VERSION : 0.1
   VAR_INPUT
      "BUFFER STATE" : Int;
      "ITEMS COUNT" : Int;
      "DOWN ELEVATOR LEFT SENSOR" : Bool;
      "BRIDGE SENSOR 1" : Bool;
      "BRIDGE SENSOR 2" : Bool;
   END_VAR
   VAR_OUTPUT
      "Z3-1 BRIDGE" : Bool;
      "Z3-2 BRIDGE" : Bool;
      "Z3-3 BRIDGE" : Bool;
   END_VAR
   VAR
      F_TRIG_Instance : F_TRIG;
      "DOWN SENSOR TRIG" : Bool;
      "BRIDGE SENSOR 1 TRIG" : Bool;
      "BRIDGE SENSOR 2 TRIG" : Bool;
      F_TRIG_BS1 : F_TRIG;
      F_TRIG_BS2 : F_TRIG;
   END_VAR
BEGIN
   #F_TRIG_Instance(CLK := #"DOWN ELEVATOR LEFT SENSOR",
                    Q => #"DOWN SENSOR TRIG");
   #F_TRIG_BS1(CLK := #"BRIDGE SENSOR 1",
               Q => #"BRIDGE SENSOR 1 TRIG");
   #F_TRIG_BS2(CLK := #"BRIDGE SENSOR 2",
               Q => #"BRIDGE SENSOR 2 TRIG");
   CASE #"ITEMS COUNT" OF
       1..2:
           #"Z3-3 BRIDGE" := 1;
           #"Z3-2 BRIDGE" := 0;
           #"Z3-3 BRIDGE" := 0;

           IF #"DOWN SENSOR TRIG" THEN
               #"Z3-3 BRIDGE" := 0;
               #"Z3-2 BRIDGE" := 0;
               #"Z3-3 BRIDGE" := 0;


           END_IF;
       3..4:
           #"Z3-3 BRIDGE" := 1;
           #"Z3-2 BRIDGE" := 1;
           #"Z3-3 BRIDGE" := 0;

           IF #"BRIDGE SENSOR 2 TRIG" AND #"DOWN SENSOR TRIG" THEN
               #"Z3-3 BRIDGE" := 0;
               #"Z3-2 BRIDGE" := 0;
               #"Z3-3 BRIDGE" := 0;

           END_IF;
       5..6:
           #"Z3-3 BRIDGE" := 1;
           #"Z3-2 BRIDGE" := 1;
           #"Z3-3 BRIDGE":=1;

           IF #"BRIDGE SENSOR 2 TRIG" AND #"DOWN SENSOR TRIG" AND #"BRIDGE SENSOR 1 TRIG" THEN
               #"Z3-3 BRIDGE" := 0;
               #"Z3-2 BRIDGE" := 0;
               #"Z3-3 BRIDGE" := 0;

           END_IF;
       ELSE 
           #"Z3-3 BRIDGE" := 0;
           #"Z3-2 BRIDGE" := 0;
           #"Z3-3 BRIDGE" := 0;

   END_CASE;
END_FUNCTION_BLOCK

FUNCTION_BLOCK "ZONE 3 ELEVATORS LOGIC"   // FB11, SCL
{ S7_Optimized_Access := 'TRUE' }
VERSION : 0.1
   VAR_INPUT
      "BUFFER STATE" : Int;
   END_VAR
   VAR_OUTPUT
      "UP ELEVATOR" : Bool;
      "DOWN ELEVATOR" : Bool;
   END_VAR
BEGIN
   IF #"BUFFER STATE" = 10 OR #"BUFFER STATE" = 33 OR #"BUFFER STATE" = 36 OR #"BUFFER STATE" = 39 THEN
       #"UP ELEVATOR" := 1;
       #"DOWN ELEVATOR" := 0;
   ELSIF #"BUFFER STATE" = 70 OR #"BUFFER STATE"=50 THEN
       #"UP ELEVATOR" := 0;
       #"DOWN ELEVATOR" := 1;
   ELSE
       #"UP ELEVATOR" := 0;
       #"DOWN ELEVATOR" := 0;
   END_IF;
END_FUNCTION_BLOCK

FUNCTION_BLOCK "ZONE 3 BRIDGE CONVS LOGIC"   // FB12, SCL
{ S7_Optimized_Access := 'TRUE' }
VERSION : 0.1
   VAR_INPUT
      "BUFFER STATE" : Int;
      "BRIDGE SENSOR 1" : Bool;
      "BRIDGE SENSOR 2" : Bool;
      "UP ELEVATOR SENSOR RIGHT" : Bool;
      "DOWN ELEVATOR LEFT SENSOR" : Bool;
      "ITEMS COUNT" : Int;
   END_VAR
   VAR_OUTPUT
      "Z3-1 BRIDGE" : Bool;
      "Z3-2 BRIDGE" : Bool;
      "Z3-3 BRIDGE" : Bool;
      "STATE 50 DONE" : Bool;
      "STATE 30 DONE" : Bool;
   END_VAR
   VAR
      "bridge sensor 1 set" : Bool;
      "bridge sensor 2 set" : Bool;
      "elevator sensor set" : Bool;
   END_VAR
BEGIN
   IF #"BUFFER STATE" = 33 THEN
       #"Z3-1 BRIDGE" := 1;
       #"Z3-2 BRIDGE" := 1;
       #"Z3-3 BRIDGE" := 1;
       IF #"BRIDGE SENSOR 2" THEN
           #"Z3-1 BRIDGE" := 0;
           #"Z3-2 BRIDGE" := 0;
           #"Z3-3 BRIDGE" := 0;
           #"STATE 30 DONE" := 1;
       END_IF;
   ELSIF #"BUFFER STATE" = 36 THEN
       #"Z3-1 BRIDGE" := 1;
       #"Z3-2 BRIDGE" := 1;
       #"Z3-3 BRIDGE" := 0;
       IF #"BRIDGE SENSOR 1" THEN
           #"Z3-1 BRIDGE" := 0;
           #"Z3-2 BRIDGE" := 0;
           #"Z3-3 BRIDGE" := 0;
           #"STATE 30 DONE" := 1;
       END_IF;
   ELSIF #"BUFFER STATE" = 39 THEN
       #"Z3-1 BRIDGE" := 1;
       #"Z3-2 BRIDGE" := 0;
       #"Z3-3 BRIDGE" := 0;
       IF #"UP ELEVATOR SENSOR RIGHT" THEN
           #"Z3-1 BRIDGE" := 0;
           #"Z3-2 BRIDGE" := 0;
           #"Z3-3 BRIDGE" := 0;
           #"STATE 30 DONE" := 1;
       END_IF;
   ELSIF #"BUFFER STATE" = 50 THEN
       CASE #"ITEMS COUNT" OF
           0..1:(*

        modified the item count to be less by one because at the cycle scan it is degreesed before it reads the current value
   *)
               #"Z3-3 BRIDGE" := 1;
               #"Z3-2 BRIDGE" := 0;
               #"Z3-1 BRIDGE" := 0;

               IF #"DOWN ELEVATOR LEFT SENSOR" THEN
                   #"Z3-3 BRIDGE" := 0;
                   #"Z3-2 BRIDGE" := 0;
                   #"Z3-1 BRIDGE" := 0;
                   #"STATE 50 DONE" := 1;

               END_IF;
           2..3:
               #"Z3-3 BRIDGE" := 1;
               #"Z3-2 BRIDGE" := 1;
               #"Z3-1 BRIDGE" := 0;

               IF #"BRIDGE SENSOR 2" THEN
                   #"bridge sensor 2 set" := 1;
               END_IF;
               IF #"DOWN ELEVATOR LEFT SENSOR" THEN
                   #"elevator sensor set" := 1;
               END_IF;
               IF #"bridge sensor 2 set" AND #"elevator sensor set" THEN
                   #"Z3-3 BRIDGE" := 0;
                   #"Z3-2 BRIDGE" := 0;
                   #"Z3-1 BRIDGE" := 0;
                   #"STATE 50 DONE" := 1;
                   #"bridge sensor 2 set" :=0;
                   #"elevator sensor set" :=0;
               END_IF;
           4..6:
               #"Z3-3 BRIDGE" := 1;
               #"Z3-2 BRIDGE" := 1;
               #"Z3-1 BRIDGE" := 1;

               IF #"BRIDGE SENSOR 2" THEN
                   #"bridge sensor 2 set" := 1;
               END_IF;
               IF #"DOWN ELEVATOR LEFT SENSOR" THEN
                   #"elevator sensor set" := 1;
               END_IF;
               IF #"BRIDGE SENSOR 1" THEN
                   #"bridge sensor 1 set" := 1;
               END_IF;
               IF #"bridge sensor 1 set" AND #"bridge sensor 2 set" AND #"elevator sensor set" THEN
                   #"Z3-3 BRIDGE" := 0;
                   #"Z3-2 BRIDGE" := 0;
                   #"Z3-1 BRIDGE" := 0;
                   #"STATE 50 DONE" := 1;
                   #"bridge sensor 2 set" := 0;
                   #"elevator sensor set" := 0;
                   #"bridge sensor 1 set" := 0;
               END_IF;
           ELSE
               #"Z3-3 BRIDGE" := 0;
               #"Z3-2 BRIDGE" := 0;
               #"Z3-1 BRIDGE" := 0;

       END_CASE;
   ELSE
       #"Z3-1 BRIDGE" := 0;
       #"Z3-2 BRIDGE" := 0;
       #"Z3-3 BRIDGE" := 0;
       #"STATE 30 DONE" := 0;
       #"STATE 50 DONE" := 0;
   END_IF;
END_FUNCTION_BLOCK

(* ===== HMI "HMI_RT_1" =====
system functions are stored by id; their names below are inferred from use
connection "HMI_Connection_1": ETHERNET, SMART_S7_1200_OMS

HMI tags "Default tag table"
   "Tag_ScreenNumber" : UInt, internal
   "DB_RackMemory_In_Production" : Int = PLC DB_RackMemory.In_Production, 1 s
   "ZONE-3 BUFFER_A_DB_BUFFER_ITEMS_COUNT_CV" : Int = PLC "ZONE-3 BUFFER_A_DB".BUFFER_ITEMS_COUNT.CV, 1 s
   "Zone_3_FB_DB_ZONE-3 BUFFER B_BUFFER_ITEMS_COUNT_CV" : Int = PLC Zone_3_FB_DB."ZONE-3 BUFFER B".BUFFER_ITEMS_COUNT.CV, 1 s
   "DB_RackMemory_SpacesOccupied" : Int = PLC DB_RackMemory.SpacesOccupied, 1 s
   "DB_HMI_Z3 BUFFER A STATUS" : Int = PLC DB_HMI."Z3 BUFFER A STATUS", 1 s
   "DB_HMI_Z1 STATUS" : Int = PLC DB_HMI."Z1 STATUS", 1 s
   "DB_HMI_Z2 STATUS" : Int = PLC DB_HMI."Z2 STATUS", 1 s
   "DB_HMI_Z3 BUFFER B STATUS" : Int = PLC DB_HMI."Z3 BUFFER B STATUS", 1 s
   "DB_HMI_Z3 ASSEMPLER STATUS" : Int = PLC DB_HMI."Z3 ASSEMPLER STATUS", 1 s
   "DB_HMI_Z5 STATUS" : Int = PLC DB_HMI."Z5 STATUS", 1 s
   "DB_HMI_Z4 UPPER STATUS" : Int = PLC DB_HMI."Z4 UPPER STATUS", 1 s
   "DB_HMI_Z4 LOWER STATUS" : Int = PLC DB_HMI."Z4 LOWER STATUS", 1 s
   "DB_HMI_FACTORY STATUS" : Int = PLC DB_HMI."FACTORY STATUS", 1 s
   "DB_RackMemory_QUANTITY TO RETRIEVE" : Int = PLC DB_RackMemory."QUANTITY TO RETRIEVE", 1 s
   "DB_RackMemory_TOTAL ORDERS" : Int = PLC DB_RackMemory."TOTAL ORDERS", 1 s
   "DB_RackMemory_TOTAL DLIEVERED" : Int = PLC DB_RackMemory."TOTAL DLIEVERED", 1 s
   "DB_RackMemory_REQUIRED QUANTITY" : Int = PLC DB_RackMemory."REQUIRED QUANTITY", 1 s
   "DB_HMI_CREATE ORDER" : Bool = PLC DB_HMI."CREATE ORDER", 1 s
   "DB_HMI_CANCEL ORDER" : Bool = PLC DB_HMI."CANCEL ORDER", 1 s
   "DB_RackMemory_FREE SPACES" : Int = PLC DB_RackMemory."FREE SPACES", 1 s
   "DB_RackMemory_Rack{1}_occupied" : Bool = PLC DB_RackMemory.Rack[1].occupied, 1 s
   "DB_RackMemory_Rack{2}_occupied" : Bool = PLC DB_RackMemory.Rack[2].occupied, 1 s
   "DB_RackMemory_Rack{3}_occupied" : Bool = PLC DB_RackMemory.Rack[3].occupied, 1 s
   "DB_RackMemory_Rack{4}_occupied" : Bool = PLC DB_RackMemory.Rack[4].occupied, 1 s
   "DB_RackMemory_Rack{5}_occupied" : Bool = PLC DB_RackMemory.Rack[5].occupied, 1 s
   "DB_RackMemory_Rack{6}_occupied" : Bool = PLC DB_RackMemory.Rack[6].occupied, 1 s
   "DB_RackMemory_Rack{7}_occupied" : Bool = PLC DB_RackMemory.Rack[7].occupied, 1 s
   "DB_RackMemory_Rack{8}_occupied" : Bool = PLC DB_RackMemory.Rack[8].occupied, 1 s
   "DB_RackMemory_Rack{9}_occupied" : Bool = PLC DB_RackMemory.Rack[9].occupied, 1 s
   "DB_RackMemory_Rack{10}_occupied" : Bool = PLC DB_RackMemory.Rack[10].occupied, 1 s
   "DB_RackMemory_Rack{11}_occupied" : Bool = PLC DB_RackMemory.Rack[11].occupied, 1 s
   "DB_RackMemory_Rack{12}_occupied" : Bool = PLC DB_RackMemory.Rack[12].occupied, 1 s
   "DB_RackMemory_Rack{13}_occupied" : Bool = PLC DB_RackMemory.Rack[13].occupied, 1 s
   "DB_RackMemory_Rack{14}_occupied" : Bool = PLC DB_RackMemory.Rack[14].occupied, 1 s
   "DB_RackMemory_Rack{15}_occupied" : Bool = PLC DB_RackMemory.Rack[15].occupied, 1 s
   "DB_RackMemory_Rack{16}_occupied" : Bool = PLC DB_RackMemory.Rack[16].occupied, 1 s
   "DB_RackMemory_Rack{17}_occupied" : Bool = PLC DB_RackMemory.Rack[17].occupied, 1 s
   "DB_RackMemory_Rack{18}_occupied" : Bool = PLC DB_RackMemory.Rack[18].occupied, 1 s
   "DB_RackMemory_Rack{19}_occupied" : Bool = PLC DB_RackMemory.Rack[19].occupied, 1 s
   "DB_RackMemory_Rack{20}_occupied" : Bool = PLC DB_RackMemory.Rack[20].occupied, 1 s
   "DB_RackMemory_Rack{21}_occupied" : Bool = PLC DB_RackMemory.Rack[21].occupied, 1 s
   "DB_RackMemory_Rack{22}_occupied" : Bool = PLC DB_RackMemory.Rack[22].occupied, 1 s
   "DB_RackMemory_Rack{23}_occupied" : Bool = PLC DB_RackMemory.Rack[23].occupied, 1 s
   "DB_RackMemory_Rack{24}_occupied" : Bool = PLC DB_RackMemory.Rack[24].occupied, 1 s
   "DB_RackMemory_Rack{25}_occupied" : Bool = PLC DB_RackMemory.Rack[25].occupied, 1 s
   "DB_RackMemory_Rack{26}_occupied" : Bool = PLC DB_RackMemory.Rack[26].occupied, 1 s
   "DB_RackMemory_Rack{27}_occupied" : Bool = PLC DB_RackMemory.Rack[27].occupied, 1 s
   "DB_RackMemory_Rack{28}_occupied" : Bool = PLC DB_RackMemory.Rack[28].occupied, 1 s
   "DB_RackMemory_Rack{29}_occupied" : Bool = PLC DB_RackMemory.Rack[29].occupied, 1 s
   "DB_RackMemory_Rack{30}_occupied" : Bool = PLC DB_RackMemory.Rack[30].occupied, 1 s
   "DB_RackMemory_Rack{31}_occupied" : Bool = PLC DB_RackMemory.Rack[31].occupied, 1 s
   "DB_RackMemory_Rack{32}_occupied" : Bool = PLC DB_RackMemory.Rack[32].occupied, 1 s
   "DB_RackMemory_Rack{33}_occupied" : Bool = PLC DB_RackMemory.Rack[33].occupied, 1 s
   "DB_RackMemory_Rack{34}_occupied" : Bool = PLC DB_RackMemory.Rack[34].occupied, 1 s
   "DB_RackMemory_Rack{35}_occupied" : Bool = PLC DB_RackMemory.Rack[35].occupied, 1 s
   "DB_RackMemory_Rack{36}_occupied" : Bool = PLC DB_RackMemory.Rack[36].occupied, 1 s
   "DB_RackMemory_Rack{37}_occupied" : Bool = PLC DB_RackMemory.Rack[37].occupied, 1 s
   "DB_RackMemory_Rack{38}_occupied" : Bool = PLC DB_RackMemory.Rack[38].occupied, 1 s
   "DB_RackMemory_Rack{39}_occupied" : Bool = PLC DB_RackMemory.Rack[39].occupied, 1 s
   "DB_RackMemory_Rack{40}_occupied" : Bool = PLC DB_RackMemory.Rack[40].occupied, 1 s
   "DB_RackMemory_Rack{41}_occupied" : Bool = PLC DB_RackMemory.Rack[41].occupied, 1 s
   "DB_RackMemory_Rack{42}_occupied" : Bool = PLC DB_RackMemory.Rack[42].occupied, 1 s
   "DB_RackMemory_Rack{43}_occupied" : Bool = PLC DB_RackMemory.Rack[43].occupied, 1 s
   "DB_RackMemory_Rack{44}_occupied" : Bool = PLC DB_RackMemory.Rack[44].occupied, 1 s
   "DB_RackMemory_Rack{45}_occupied" : Bool = PLC DB_RackMemory.Rack[45].occupied, 1 s
   "DB_RackMemory_Rack{46}_occupied" : Bool = PLC DB_RackMemory.Rack[46].occupied, 1 s
   "DB_RackMemory_Rack{47}_occupied" : Bool = PLC DB_RackMemory.Rack[47].occupied, 1 s
   "DB_RackMemory_Rack{48}_occupied" : Bool = PLC DB_RackMemory.Rack[48].occupied, 1 s
   "DB_RackMemory_Rack{49}_occupied" : Bool = PLC DB_RackMemory.Rack[49].occupied, 1 s
   "DB_RackMemory_Rack{50}_occupied" : Bool = PLC DB_RackMemory.Rack[50].occupied, 1 s
   "DB_RackMemory_Rack{51}_occupied" : Bool = PLC DB_RackMemory.Rack[51].occupied, 1 s
   "DB_RackMemory_Rack{52}_occupied" : Bool = PLC DB_RackMemory.Rack[52].occupied, 1 s
   "DB_RackMemory_Rack{53}_occupied" : Bool = PLC DB_RackMemory.Rack[53].occupied, 1 s
   "DB_RackMemory_Rack{54}_occupied" : Bool = PLC DB_RackMemory.Rack[54].occupied, 1 s
   "DB_RackMemory_Rack{55}_occupied" : Bool = PLC DB_RackMemory.Rack[55].occupied, 1 s
   "DB_RackMemory_Rack{56}_occupied" : Bool = PLC DB_RackMemory.Rack[56].occupied, 1 s
   "DB_RackMemory_Rack{57}_occupied" : Bool = PLC DB_RackMemory.Rack[57].occupied, 1 s
   "DB_RackMemory_Rack{58}_occupied" : Bool = PLC DB_RackMemory.Rack[58].occupied, 1 s
   "DB_RackMemory_Rack{59}_occupied" : Bool = PLC DB_RackMemory.Rack[59].occupied, 1 s
   "DB_RackMemory_Rack{60}_occupied" : Bool = PLC DB_RackMemory.Rack[60].occupied, 1 s
   "DB_RackMemory_Rack{61}_occupied" : Bool = PLC DB_RackMemory.Rack[61].occupied, 1 s
   "DB_RackMemory_Rack{62}_occupied" : Bool = PLC DB_RackMemory.Rack[62].occupied, 1 s
   "DB_RackMemory_Rack{63}_occupied" : Bool = PLC DB_RackMemory.Rack[63].occupied, 1 s
   "DB_RackMemory_Rack{64}_occupied" : Bool = PLC DB_RackMemory.Rack[64].occupied, 1 s
   "DB_RackMemory_Rack{65}_occupied" : Bool = PLC DB_RackMemory.Rack[65].occupied, 1 s
   "DB_RackMemory_Rack{66}_occupied" : Bool = PLC DB_RackMemory.Rack[66].occupied, 1 s
   "DB_RackMemory_Rack{67}_occupied" : Bool = PLC DB_RackMemory.Rack[67].occupied, 1 s
   "DB_RackMemory_Rack{68}_occupied" : Bool = PLC DB_RackMemory.Rack[68].occupied, 1 s
   "DB_RackMemory_Rack{69}_occupied" : Bool = PLC DB_RackMemory.Rack[69].occupied, 1 s
   "DB_RackMemory_Rack{70}_occupied" : Bool = PLC DB_RackMemory.Rack[70].occupied, 1 s
   "DB_RackMemory_Rack{71}_occupied" : Bool = PLC DB_RackMemory.Rack[71].occupied, 1 s
   "DB_RackMemory_Rack{72}_occupied" : Bool = PLC DB_RackMemory.Rack[72].occupied, 1 s
   "DB_RackMemory_Rack{73}_occupied" : Bool = PLC DB_RackMemory.Rack[73].occupied, 1 s
   "DB_RackMemory_Rack{74}_occupied" : Bool = PLC DB_RackMemory.Rack[74].occupied, 1 s
   "DB_RackMemory_Rack{75}_occupied" : Bool = PLC DB_RackMemory.Rack[75].occupied, 1 s
   "DB_RackMemory_Rack{76}_occupied" : Bool = PLC DB_RackMemory.Rack[76].occupied, 1 s
   "DB_RackMemory_Rack{77}_occupied" : Bool = PLC DB_RackMemory.Rack[77].occupied, 1 s
   "DB_RackMemory_Rack{78}_occupied" : Bool = PLC DB_RackMemory.Rack[78].occupied, 1 s
   "DB_RackMemory_Rack{79}_occupied" : Bool = PLC DB_RackMemory.Rack[79].occupied, 1 s
   "DB_RackMemory_Rack{80}_occupied" : Bool = PLC DB_RackMemory.Rack[80].occupied, 1 s
   "DB_RackMemory_Rack{81}_occupied" : Bool = PLC DB_RackMemory.Rack[81].occupied, 1 s
   "DB_RackMemory_Rack{82}_occupied" : Bool = PLC DB_RackMemory.Rack[82].occupied, 1 s
   "DB_RackMemory_Rack{83}_occupied" : Bool = PLC DB_RackMemory.Rack[83].occupied, 1 s
   "DB_RackMemory_Rack{84}_occupied" : Bool = PLC DB_RackMemory.Rack[84].occupied, 1 s
   "DB_RackMemory_Rack{85}_occupied" : Bool = PLC DB_RackMemory.Rack[85].occupied, 1 s
   "DB_RackMemory_Rack{86}_occupied" : Bool = PLC DB_RackMemory.Rack[86].occupied, 1 s
   "DB_RackMemory_Rack{87}_occupied" : Bool = PLC DB_RackMemory.Rack[87].occupied, 1 s
   "DB_RackMemory_Rack{88}_occupied" : Bool = PLC DB_RackMemory.Rack[88].occupied, 1 s
   "DB_RackMemory_Rack{89}_occupied" : Bool = PLC DB_RackMemory.Rack[89].occupied, 1 s
   "DB_RackMemory_Rack{90}_occupied" : Bool = PLC DB_RackMemory.Rack[90].occupied, 1 s
   "DB_RackMemory_Rack{91}_occupied" : Bool = PLC DB_RackMemory.Rack[91].occupied, 1 s
   "DB_RackMemory_Rack{92}_occupied" : Bool = PLC DB_RackMemory.Rack[92].occupied, 1 s
   "DB_RackMemory_Rack{93}_occupied" : Bool = PLC DB_RackMemory.Rack[93].occupied, 1 s
   "DB_RackMemory_Rack{94}_occupied" : Bool = PLC DB_RackMemory.Rack[94].occupied, 1 s
   "DB_RackMemory_Rack{95}_occupied" : Bool = PLC DB_RackMemory.Rack[95].occupied, 1 s
   "DB_RackMemory_Rack{96}_occupied" : Bool = PLC DB_RackMemory.Rack[96].occupied, 1 s
   "DB_RackMemory_Rack{97}_occupied" : Bool = PLC DB_RackMemory.Rack[97].occupied, 1 s
   "DB_RackMemory_Rack{98}_occupied" : Bool = PLC DB_RackMemory.Rack[98].occupied, 1 s
   "DB_RackMemory_Rack{99}_occupied" : Bool = PLC DB_RackMemory.Rack[99].occupied, 1 s
   "DB_RackMemory_Rack{100}_occupied" : Bool = PLC DB_RackMemory.Rack[100].occupied, 1 s
   "DB_RackMemory_Rack{101}_occupied" : Bool = PLC DB_RackMemory.Rack[101].occupied, 1 s
   "DB_RackMemory_Rack{102}_occupied" : Bool = PLC DB_RackMemory.Rack[102].occupied, 1 s
   "DB_RackMemory_Rack{103}_occupied" : Bool = PLC DB_RackMemory.Rack[103].occupied, 1 s
   "DB_RackMemory_Rack{104}_occupied" : Bool = PLC DB_RackMemory.Rack[104].occupied, 1 s
   "DB_RackMemory_Rack{105}_occupied" : Bool = PLC DB_RackMemory.Rack[105].occupied, 1 s
   "DB_RackMemory_Rack{106}_occupied" : Bool = PLC DB_RackMemory.Rack[106].occupied, 1 s
   "DB_RackMemory_Rack{107}_occupied" : Bool = PLC DB_RackMemory.Rack[107].occupied, 1 s
   "DB_RackMemory_Rack{108}_occupied" : Bool = PLC DB_RackMemory.Rack[108].occupied, 1 s
   "DB_HMI_CRANE TARGET" : Int = PLC DB_HMI."CRANE TARGET", 1 s
   "DB_HMI_CRANE SIDE" : Int = PLC DB_HMI."CRANE SIDE", 1 s
   "DB_HMI_ASSEMPLER X" : Real = PLC DB_HMI."ASSEMPLER X", 1 s
   "DB_HMI_ASSEMPLER Z" : Real = PLC DB_HMI."ASSEMPLER Z", 1 s
   "DB_RackMemory_ReckMemoryReset" : Bool = PLC DB_RackMemory.ReckMemoryReset, 1 s
   "DB_RackMemory_InProductionReset" : Bool = PLC DB_RackMemory.InProductionReset, 1 s
   "DB_HMI_CRANE LIFT" : Bool = PLC DB_HMI."CRANE LIFT", 1 s
   "DB_HMI_CRANE LEFT" : Bool = PLC DB_HMI."CRANE LEFT", 1 s
   "DB_HMI_CRANE RIGHT" : Bool = PLC DB_HMI."CRANE RIGHT", 1 s
   "DB_HMI_ASSEMPLER ROT CW" : Bool = PLC DB_HMI."ASSEMPLER ROT CW", 1 s
   "DB_HMI_ASSEMPLER ROT CCW" : Bool = PLC DB_HMI."ASSEMPLER ROT CCW", 1 s
   "DB_HMI_ASSEMPLER GRAB" : Bool = PLC DB_HMI."ASSEMPLER GRAB", 1 s
   "DB_RackMemory_RETRIEVE" : Bool = PLC DB_RackMemory.RETRIEVE, 1 s
   "CURRENT USER" : WString[254] AT %DB1.DBX0.0
   "DB_HMI_MAINTENANCE MODE" : Bool = PLC DB_HMI."MAINTENANCE MODE", 1 s

HMI tags "Alarm tag table"
   "Alarm_Trigger" : Word = PLC Alarm_trigger AT %MW100, 1 s

discrete alarms
   1: 'Emergency button is pressed', class Errors, trigger "Alarm_Trigger" bit 0
   2: 'MACHINE A HAS AN ERROR AND STOPPED WORKING', class Errors, trigger "Alarm_Trigger" bit 1
   3: 'MACHINE B HAS AN ERROR AND STOPPED WORKING', class Errors, trigger "Alarm_Trigger" bit 2
   4: 'BUFFER A HAS A PROBLEM AND STOPPED RESPONDING', class Errors, trigger "Alarm_Trigger" bit 3
   5: 'BUFFER B HAS A PROBLEM AND STOPPED WORKING', class Errors, trigger "Alarm_Trigger" bit 4
   6: 'ASSEMPLER HAS A PROBLEM AND STOPPED RESPONDING', class Errors, trigger "Alarm_Trigger" bit 5
   7: 'PALLETIZER HAS A PROBLEM AND STOPPED RESPONDING', class Errors, trigger "Alarm_Trigger" bit 6
   8: 'CRANE HAS A PROBLEM AND STOPPED RESPONDING', class Errors, trigger "Alarm_Trigger" bit 7

Template "Template_1" 800x480
   Button "Template_Button" at 714,429 size 71x50; TextOff 'Text'
   Button "Template_Button_1" at 614,429 size 71x50; TextOff 'Text'
   Button "Template_Button_2" at 514,429 size 71x50; TextOff 'Text'
   Button "Template_Button_3" at 414,429 size 71x50; TextOff 'Text'
   Button "Template_Button_4" at 314,429 size 71x50; TextOff 'Text'
   Button "Template_Button_5" at 214,429 size 71x50; TextOff 'Text'
   Button "Template_Button_6" at 114,429 size 71x50; TextOff 'Text'
   Button "Template_Button_7" at 14,429 size 71x50; TextOff 'Text'
   SymbolicIOField "Symbolic_IO_Field_Screen" at 93,9 size 600x33; TextOff '0'; TextOn '1'; TextList "TextList_ScreenNames"
      ProcessValue <- "Tag_ScreenNumber"
      on Change: ActivateScreenByNumber("Tag_ScreenNumber", 0)
   DateTimeField "HmiScreenItemData" at 695,25 size 105x25
   DateTimeField "HmiScreenItemData_1" at 695,0 size 105x25
   GraphicView "Logo" at 0,0 size 91x51; Picture "Logo of HMI_1"

screen "Production" 800x480
   Button "Button_12" at 69,415 size 163x52; TextOff 'Overview'
      on Release: ActivateScreen("Overview", 0)
   Button "Button_13" at 238,415 size 163x52; TextOff 'Warehouse'
      on Release: ActivateScreen("Warehouse", 0)
   Button "Button_14" at 408,415 size 163x52; TextOff 'Alarms'
      on Release: ActivateScreen("Alarms", 0)
   Button "Button_15" at 578,415 size 163x52; TextOff 'Maintenance'; Authorization "Maintenance"
      on Release: ActivateScreen("Maintenance", 0)
   TextField "Text field_1" at 310,0 size 180x44; Text 'Production'
   TextField "Text field_2" at 12,130 size 86x23; Text 'Quantity :'
   IOField "I/O field_1" at 124,121 size 96x32; Authorization "Operate"; FormatPattern 99
      ProcessValue <- "DB_RackMemory_QUANTITY TO RETRIEVE"
   Button "Button_1" at 65,221 size 96x32; TextOff 'Order'; Authorization "Operate"
      on Press: SetBit("DB_RackMemory_RETRIEVE")
   TextField "Text field_3" at 128,307 size 97x23; Text 'In Storage:'
   TextField "Text field_4" at 381,307 size 164x23; Text 'In Production lines:'
   IOField "I/O field_2" at 255,298 size 96x32; FormatPattern 999
      ProcessValue <- "DB_RackMemory_SpacesOccupied"
   IOField "I/O field_3" at 575,298 size 96x32; FormatPattern 99
      ProcessValue <- "DB_RackMemory_In_Production"
   TextField "Text field_5" at 27,70 size 163x33; Text 'Create Order:'
   TextField "Text field_6" at 312,70 size 175x33; Text 'Current Order:'
   TextField "Text field_7" at 247,130 size 161x23; Text 'Required Products:'
   TextField "Text field_8" at 240,183 size 174x23; Text 'Products Remaining:'
   TextField "Text field_9" at 610,70 size 124x33; Text 'Summary:'
   TextField "Text field_10" at 558,130 size 113x23; Text 'Total Orders:'
   TextField "Text field_11" at 537,183 size 147x23; Text 'Total Delievered:'
   Button "Button_2" at 352,221 size 96x32; TextOff 'Cancel'; Authorization "Operate"
      on Press: SetBit("DB_HMI_CANCEL ORDER")
      on Release: ResetBit("DB_HMI_CANCEL ORDER")
   IOField "I/O field_4" at 425,121 size 96x32; FormatPattern 99
      ProcessValue <- "DB_RackMemory_REQUIRED QUANTITY"
   IOField "I/O field_5" at 425,174 size 96x32; FormatPattern 99
      ProcessValue <- "DB_RackMemory_QUANTITY TO RETRIEVE"
   IOField "I/O field_6" at 690,121 size 96x32; FormatPattern 999
      ProcessValue <- "DB_RackMemory_TOTAL ORDERS"
   IOField "I/O field_7" at 690,174 size 96x32; FormatPattern 999
      ProcessValue <- "DB_RackMemory_TOTAL DLIEVERED"
   Button "Button_3" at 11,10 size 96x32; TextOff 'LOG IN'
      on Release: function_f41c6f6c("CURRENT USER")
      on Press: function_a2a04561()
   Button "Button_4" at 126,8 size 96x32; TextOff 'LOG OUT'
      on Press: function_f23ef4c9(); SetTag("CURRENT USER", '""')
   IOField "I/O field_13" at 685,3 size 106x32; FormatPattern ??????????????????????????????????????????????????????????????????????
      ProcessValue <- "CURRENT USER"
   TextField "Text field_12" at 542,8 size 140x23; Text 'CURRENT USER:'

screen "Warehouse" 800x480
   Rectangle "Rectangle_1" at 698,216 size 20x20
      Appearance <- "DB_RackMemory_Rack{1}_occupied"
   Rectangle "Rectangle_2" at 678,216 size 20x20
      Appearance <- "DB_RackMemory_Rack{2}_occupied"
   Rectangle "Rectangle_3" at 658,216 size 20x20
      Appearance <- "DB_RackMemory_Rack{3}_occupied"
   Rectangle "Rectangle_4" at 638,216 size 20x20
      Appearance <- "DB_RackMemory_Rack{4}_occupied"
   Rectangle "Rectangle_5" at 618,216 size 20x20
      Appearance <- "DB_RackMemory_Rack{5}_occupied"
   Rectangle "Rectangle_6" at 598,216 size 20x20
      Appearance <- "DB_RackMemory_Rack{6}_occupied"
   Rectangle "Rectangle_7" at 578,216 size 20x20
      Appearance <- "DB_RackMemory_Rack{7}_occupied"
   Rectangle "Rectangle_8" at 558,216 size 20x20
      Appearance <- "DB_RackMemory_Rack{8}_occupied"
   Rectangle "Rectangle_9" at 538,216 size 20x20
      Appearance <- "DB_RackMemory_Rack{9}_occupied"
   Rectangle "Rectangle_10" at 698,196 size 20x20
      Appearance <- "DB_RackMemory_Rack{10}_occupied"
   Rectangle "Rectangle_11" at 678,196 size 20x20
      Appearance <- "DB_RackMemory_Rack{11}_occupied"
   Rectangle "Rectangle_12" at 658,196 size 20x20
      Appearance <- "DB_RackMemory_Rack{12}_occupied"
   Rectangle "Rectangle_13" at 638,196 size 20x20
      Appearance <- "DB_RackMemory_Rack{13}_occupied"
   Rectangle "Rectangle_14" at 618,196 size 20x20
      Appearance <- "DB_RackMemory_Rack{14}_occupied"
   Rectangle "Rectangle_15" at 598,196 size 20x20
      Appearance <- "DB_RackMemory_Rack{15}_occupied"
   Rectangle "Rectangle_16" at 578,196 size 20x20
      Appearance <- "DB_RackMemory_Rack{16}_occupied"
   Rectangle "Rectangle_17" at 558,196 size 20x20
      Appearance <- "DB_RackMemory_Rack{17}_occupied"
   Rectangle "Rectangle_18" at 538,196 size 20x20
      Appearance <- "DB_RackMemory_Rack{18}_occupied"
   Rectangle "Rectangle_19" at 698,176 size 20x20
      Appearance <- "DB_RackMemory_Rack{19}_occupied"
   Rectangle "Rectangle_20" at 678,176 size 20x20
      Appearance <- "DB_RackMemory_Rack{20}_occupied"
   Rectangle "Rectangle_21" at 658,176 size 20x20
      Appearance <- "DB_RackMemory_Rack{21}_occupied"
   Rectangle "Rectangle_22" at 638,176 size 20x20
      Appearance <- "DB_RackMemory_Rack{22}_occupied"
   Rectangle "Rectangle_23" at 618,176 size 20x20
      Appearance <- "DB_RackMemory_Rack{23}_occupied"
   Rectangle "Rectangle_24" at 598,176 size 20x20
      Appearance <- "DB_RackMemory_Rack{24}_occupied"
   Rectangle "Rectangle_25" at 578,176 size 20x20
      Appearance <- "DB_RackMemory_Rack{25}_occupied"
   Rectangle "Rectangle_26" at 558,176 size 20x20
      Appearance <- "DB_RackMemory_Rack{26}_occupied"
   Rectangle "Rectangle_27" at 538,176 size 20x20
      Appearance <- "DB_RackMemory_Rack{27}_occupied"
   Rectangle "Rectangle_28" at 698,156 size 20x20
      Appearance <- "DB_RackMemory_Rack{28}_occupied"
   Rectangle "Rectangle_29" at 678,156 size 20x20
      Appearance <- "DB_RackMemory_Rack{29}_occupied"
   Rectangle "Rectangle_30" at 658,156 size 20x20
      Appearance <- "DB_RackMemory_Rack{30}_occupied"
   Rectangle "Rectangle_31" at 638,156 size 20x20
      Appearance <- "DB_RackMemory_Rack{31}_occupied"
   Rectangle "Rectangle_32" at 618,156 size 20x20
      Appearance <- "DB_RackMemory_Rack{32}_occupied"
   Rectangle "Rectangle_33" at 598,156 size 20x20
      Appearance <- "DB_RackMemory_Rack{33}_occupied"
   Rectangle "Rectangle_34" at 578,156 size 20x20
      Appearance <- "DB_RackMemory_Rack{34}_occupied"
   Rectangle "Rectangle_35" at 558,156 size 20x20
      Appearance <- "DB_RackMemory_Rack{35}_occupied"
   Rectangle "Rectangle_36" at 538,156 size 20x20
      Appearance <- "DB_RackMemory_Rack{36}_occupied"
   Rectangle "Rectangle_37" at 698,136 size 20x20
      Appearance <- "DB_RackMemory_Rack{37}_occupied"
   Rectangle "Rectangle_38" at 678,136 size 20x20
      Appearance <- "DB_RackMemory_Rack{38}_occupied"
   Rectangle "Rectangle_39" at 658,136 size 20x20
      Appearance <- "DB_RackMemory_Rack{39}_occupied"
   Rectangle "Rectangle_40" at 638,136 size 20x20
      Appearance <- "DB_RackMemory_Rack{40}_occupied"
   Rectangle "Rectangle_41" at 618,136 size 20x20
      Appearance <- "DB_RackMemory_Rack{41}_occupied"
   Rectangle "Rectangle_42" at 598,136 size 20x20
      Appearance <- "DB_RackMemory_Rack{42}_occupied"
   Rectangle "Rectangle_43" at 578,136 size 20x20
      Appearance <- "DB_RackMemory_Rack{43}_occupied"
   Rectangle "Rectangle_44" at 558,136 size 20x20
      Appearance <- "DB_RackMemory_Rack{44}_occupied"
   Rectangle "Rectangle_45" at 538,136 size 20x20
      Appearance <- "DB_RackMemory_Rack{45}_occupied"
   Rectangle "Rectangle_46" at 698,116 size 20x20
      Appearance <- "DB_RackMemory_Rack{46}_occupied"
   Rectangle "Rectangle_47" at 678,116 size 20x20
      Appearance <- "DB_RackMemory_Rack{47}_occupied"
   Rectangle "Rectangle_48" at 658,116 size 20x20
      Appearance <- "DB_RackMemory_Rack{48}_occupied"
   Rectangle "Rectangle_49" at 638,116 size 20x20
      Appearance <- "DB_RackMemory_Rack{49}_occupied"
   Rectangle "Rectangle_50" at 618,116 size 20x20
      Appearance <- "DB_RackMemory_Rack{50}_occupied"
   Rectangle "Rectangle_51" at 598,116 size 20x20
      Appearance <- "DB_RackMemory_Rack{51}_occupied"
   Rectangle "Rectangle_52" at 578,116 size 20x20
      Appearance <- "DB_RackMemory_Rack{52}_occupied"
   Rectangle "Rectangle_53" at 558,116 size 20x20
      Appearance <- "DB_RackMemory_Rack{53}_occupied"
   Rectangle "Rectangle_54" at 538,116 size 20x20
      Appearance <- "DB_RackMemory_Rack{54}_occupied"
   Rectangle "Rectangle_69" at 142,196 size 20x20
      Appearance <- "DB_RackMemory_Rack{69}_occupied"
   Rectangle "Rectangle_55" at 242,216 size 20x20
      Appearance <- "DB_RackMemory_Rack{55}_occupied"
   Rectangle "Rectangle_56" at 222,216 size 20x20
      Appearance <- "DB_RackMemory_Rack{56}_occupied"
   Rectangle "Rectangle_57" at 202,216 size 20x20
      Appearance <- "DB_RackMemory_Rack{57}_occupied"
   Rectangle "Rectangle_58" at 182,216 size 20x20
      Appearance <- "DB_RackMemory_Rack{58}_occupied"
   Rectangle "Rectangle_59" at 162,216 size 20x20
      Appearance <- "DB_RackMemory_Rack{59}_occupied"
   Rectangle "Rectangle_60" at 142,216 size 20x20
      Appearance <- "DB_RackMemory_Rack{60}_occupied"
   Rectangle "Rectangle_61" at 122,216 size 20x20
      Appearance <- "DB_RackMemory_Rack{61}_occupied"
   Rectangle "Rectangle_62" at 102,216 size 20x20
      Appearance <- "DB_RackMemory_Rack{62}_occupied"
   Rectangle "Rectangle_63" at 82,216 size 20x20
      Appearance <- "DB_RackMemory_Rack{63}_occupied"
   Rectangle "Rectangle_64" at 242,196 size 20x20
      Appearance <- "DB_RackMemory_Rack{64}_occupied"
   Rectangle "Rectangle_65" at 222,196 size 20x20
      Appearance <- "DB_RackMemory_Rack{65}_occupied"
   Rectangle "Rectangle_66" at 202,196 size 20x20
      Appearance <- "DB_RackMemory_Rack{66}_occupied"
   Rectangle "Rectangle_67" at 182,196 size 20x20
      Appearance <- "DB_RackMemory_Rack{67}_occupied"
   Rectangle "Rectangle_68" at 162,196 size 20x20
      Appearance <- "DB_RackMemory_Rack{68}_occupied"
   Rectangle "Rectangle_70" at 122,196 size 20x20
      Appearance <- "DB_RackMemory_Rack{70}_occupied"
   Rectangle "Rectangle_71" at 102,196 size 20x20
      Appearance <- "DB_RackMemory_Rack{71}_occupied"
   Rectangle "Rectangle_72" at 82,196 size 20x20
      Appearance <- "DB_RackMemory_Rack{72}_occupied"
   Rectangle "Rectangle_73" at 242,176 size 20x20
      Appearance <- "DB_RackMemory_Rack{73}_occupied"
   Rectangle "Rectangle_74" at 222,176 size 20x20
      Appearance <- "DB_RackMemory_Rack{74}_occupied"
   Rectangle "Rectangle_75" at 202,176 size 20x20
      Appearance <- "DB_RackMemory_Rack{75}_occupied"
   Rectangle "Rectangle_76" at 182,176 size 20x20
      Appearance <- "DB_RackMemory_Rack{76}_occupied"
   Rectangle "Rectangle_77" at 162,176 size 20x20
      Appearance <- "DB_RackMemory_Rack{77}_occupied"
   Rectangle "Rectangle_78" at 142,176 size 20x20
      Appearance <- "DB_RackMemory_Rack{78}_occupied"
   Rectangle "Rectangle_79" at 122,176 size 20x20
      Appearance <- "DB_RackMemory_Rack{79}_occupied"
   Rectangle "Rectangle_80" at 102,176 size 20x20
      Appearance <- "DB_RackMemory_Rack{80}_occupied"
   Rectangle "Rectangle_81" at 82,176 size 20x20
      Appearance <- "DB_RackMemory_Rack{81}_occupied"
   Rectangle "Rectangle_82" at 242,156 size 20x20
      Appearance <- "DB_RackMemory_Rack{82}_occupied"
   Rectangle "Rectangle_83" at 222,156 size 20x20
      Appearance <- "DB_RackMemory_Rack{83}_occupied"
   Rectangle "Rectangle_84" at 202,156 size 20x20
      Appearance <- "DB_RackMemory_Rack{84}_occupied"
   Rectangle "Rectangle_85" at 182,156 size 20x20
      Appearance <- "DB_RackMemory_Rack{85}_occupied"
   Rectangle "Rectangle_86" at 162,156 size 20x20
      Appearance <- "DB_RackMemory_Rack{86}_occupied"
   Rectangle "Rectangle_87" at 142,156 size 20x20
      Appearance <- "DB_RackMemory_Rack{87}_occupied"
   Rectangle "Rectangle_88" at 122,156 size 20x20
      Appearance <- "DB_RackMemory_Rack{88}_occupied"
   Rectangle "Rectangle_89" at 102,156 size 20x20
      Appearance <- "DB_RackMemory_Rack{89}_occupied"
   Rectangle "Rectangle_90" at 82,156 size 20x20
      Appearance <- "DB_RackMemory_Rack{90}_occupied"
   Rectangle "Rectangle_91" at 242,136 size 20x20
      Appearance <- "DB_RackMemory_Rack{91}_occupied"
   Rectangle "Rectangle_92" at 222,136 size 20x20
      Appearance <- "DB_RackMemory_Rack{92}_occupied"
   Rectangle "Rectangle_93" at 202,136 size 20x20
      Appearance <- "DB_RackMemory_Rack{93}_occupied"
   Rectangle "Rectangle_94" at 182,136 size 20x20
      Appearance <- "DB_RackMemory_Rack{94}_occupied"
   Rectangle "Rectangle_95" at 162,136 size 20x20
      Appearance <- "DB_RackMemory_Rack{95}_occupied"
   Rectangle "Rectangle_96" at 142,136 size 20x20
      Appearance <- "DB_RackMemory_Rack{96}_occupied"
   Rectangle "Rectangle_97" at 122,136 size 20x20
      Appearance <- "DB_RackMemory_Rack{97}_occupied"
   Rectangle "Rectangle_98" at 102,136 size 20x20
      Appearance <- "DB_RackMemory_Rack{98}_occupied"
   Rectangle "Rectangle_99" at 82,136 size 20x20
      Appearance <- "DB_RackMemory_Rack{99}_occupied"
   Rectangle "Rectangle_100" at 242,116 size 20x20
      Appearance <- "DB_RackMemory_Rack{100}_occupied"
   Rectangle "Rectangle_101" at 222,116 size 20x20
      Appearance <- "DB_RackMemory_Rack{101}_occupied"
   Rectangle "Rectangle_102" at 202,116 size 20x20
      Appearance <- "DB_RackMemory_Rack{102}_occupied"
   Rectangle "Rectangle_103" at 182,116 size 20x20
      Appearance <- "DB_RackMemory_Rack{103}_occupied"
   Rectangle "Rectangle_104" at 162,116 size 20x20
      Appearance <- "DB_RackMemory_Rack{104}_occupied"
   Rectangle "Rectangle_105" at 142,116 size 20x20
      Appearance <- "DB_RackMemory_Rack{105}_occupied"
   Rectangle "Rectangle_106" at 122,116 size 20x20
      Appearance <- "DB_RackMemory_Rack{106}_occupied"
   Rectangle "Rectangle_107" at 102,116 size 20x20
      Appearance <- "DB_RackMemory_Rack{107}_occupied"
   Rectangle "Rectangle_108" at 82,116 size 20x20
      Appearance <- "DB_RackMemory_Rack{108}_occupied"
   Button "Button_12" at 69,415 size 163x52; TextOff 'Overview'
      on Release: ActivateScreen("Overview", 0)
   Button "Button_13" at 238,415 size 163x52; TextOff 'Production'; Authorization "Operate"
      on Release: ActivateScreen("Production", 0)
   Button "Button_14" at 408,415 size 163x52; TextOff 'Alarms'
      on Release: ActivateScreen("Alarms", 0)
   Button "Button_15" at 578,415 size 163x52; TextOff 'Maintenance'; Authorization "Maintenance"
      on Release: ActivateScreen("Maintenance", 0)
   TextField "Text field_1" at 304,0 size 185x44; Text 'Warehouse'
   TextField "Text field_2" at 562,77 size 132x32; Text 'Right Rack'
   TextField "Text field_3" at 115,77 size 115x32; Text 'Left Rack'
   Group "Group_1" at 538,116 size 180x120
   TextField "Text field_4" at 723,215 size 15x23; Text '1'
   TextField "Text field_5" at 506,111 size 25x23; Text '54'
   TextField "Text field_8" at 718,194 size 25x23; Text '10'
   TextField "Text field_9" at 718,173 size 25x23; Text '19'
   TextField "Text field_10" at 718,152 size 25x23; Text '28'
   TextField "Text field_11" at 718,131 size 25x23; Text '37'
   TextField "Text field_12" at 718,111 size 25x23; Text '46'
   TextField "Text field_13" at 511,217 size 15x23; Text '9'
   TextField "Text field_14" at 506,195 size 25x23; Text '18'
   TextField "Text field_15" at 506,174 size 25x23; Text '27'
   TextField "Text field_16" at 506,153 size 25x23; Text '36'
   TextField "Text field_17" at 506,132 size 25x23; Text '45'
   TextField "Text field_6" at 272,218 size 15x23; Text '1'
   TextField "Text field_7" at 267,197 size 25x23; Text '10'
   TextField "Text field_18" at 267,176 size 25x23; Text '19'
   TextField "Text field_19" at 267,155 size 25x23; Text '28'
   TextField "Text field_20" at 267,134 size 25x23; Text '37'
   TextField "Text field_21" at 267,114 size 25x23; Text '46'
   TextField "Text field_22" at 53,112 size 25x23; Text '54'
   TextField "Text field_23" at 58,218 size 15x23; Text '9'
   TextField "Text field_24" at 53,196 size 25x23; Text '18'
   TextField "Text field_25" at 53,175 size 25x23; Text '27'
   TextField "Text field_26" at 53,154 size 25x23; Text '36'
   TextField "Text field_27" at 53,133 size 25x23; Text '45'
   TextField "Text field_28" at 291,295 size 129x23; Text 'Total Capacity:'
   TextField "Text field_29" at 291,330 size 51x23; Text 'Used:'
   TextField "Text field_30" at 291,363 size 47x23; Text 'Free:'
   IOField "I/O field_2" at 423,321 size 82x32; FormatPattern 999
      ProcessValue <- "DB_RackMemory_SpacesOccupied"
   IOField "I/O field_3" at 423,358 size 83x32; FormatPattern 999
      ProcessValue <- "DB_RackMemory_FREE SPACES"
   TextField "Text field_31" at 447,295 size 35x23; Text '108'
   Group "Group" at 82,116 size 180x120
   Button "Button_1" at 11,10 size 96x32; TextOff 'LOG IN'
      on Release: function_f41c6f6c("CURRENT USER")
      on Press: function_a2a04561()
   Button "Button_2" at 126,8 size 96x32; TextOff 'LOG OUT'
      on Press: function_f23ef4c9(); SetTag("CURRENT USER", '""')
   IOField "I/O field_13" at 685,3 size 106x32; FormatPattern ??????????????????????????????????????????????????????????????????????
      ProcessValue <- "CURRENT USER"
   TextField "Text field_32" at 542,8 size 140x23; Text 'CURRENT USER:'

screen "Alarms" 800x480
   Button "Button_12" at 69,415 size 163x52; TextOff 'OverView'
      on Release: ActivateScreen("Overview", 0)
   Button "Button_13" at 238,417 size 163x52; TextOff 'Production'; Authorization "Operate"
      on Release: ActivateScreen("Production", 0)
   Button "Button_14" at 408,415 size 163x52; TextOff 'Warehouse'
      on Release: ActivateScreen("Warehouse", 0)
   Button "Button_15" at 578,415 size 163x52; TextOff 'Maintenance'; Authorization "Maintenance"
      on Release: ActivateScreen("Maintenance", 0)
   Button "Button_1" at 11,10 size 96x32; TextOff 'LOG IN'
      on Release: function_f41c6f6c("CURRENT USER")
      on Press: function_a2a04561()
   Button "Button_2" at 126,8 size 96x32; TextOff 'LOG OUT'
      on Press: function_f23ef4c9(); SetTag("CURRENT USER", '""')
   IOField "I/O field_13" at 685,3 size 106x32; FormatPattern ??????????????????????????????????????????????????????????????????????
      ProcessValue <- "CURRENT USER"
   TextField "Text field_2" at 542,8 size 153x23; Text 'CURRENT USER:'
   TextField "Text field_1" at 342,0 size 117x44; Text 'Alarms'
   AlarmView "Alarm view_1" at 0,60 size 799x210
   AlarmView "Alarm view_2" at 0,270 size 799x142

screen "Maintenance" 800x480
   Button "Button_12" at 69,415 size 163x52; TextOff 'Overview'
      on Release: ActivateScreen("Overview", 0)
   Button "Button_13" at 238,415 size 163x52; TextOff 'Production'; Authorization "Operate"
      on Release: ActivateScreen("Production", 0)
   Button "Button_14" at 408,415 size 163x52; TextOff 'Warehouse'
      on Release: ActivateScreen("Warehouse", 0)
   Button "Button_15" at 578,415 size 163x52; TextOff 'Alarms'
      on Release: ActivateScreen("Alarms", 0)
   TextField "Text field_1" at 295,0 size 210x44; Text 'Maintenance'
   TextField "Text field_2" at 45,62 size 165x32; Text 'Crane Control'
   TextField "Text field_3" at 291,62 size 218x32; Text 'Assempler Control'
   TextField "Text field_4" at 43,120 size 66x23; Text 'Target:'
   IOField "I/O field_1" at 126,111 size 96x32; Authorization "Maintenance"; FormatPattern 999
      ProcessValue <- "DB_HMI_CRANE TARGET"
   Button "Button_1" at 80,198 size 96x32; TextOff 'Lift'; Authorization "Maintenance"
      on Press: InvertBit("DB_HMI_CRANE LIFT")
      Appearance <- "DB_HMI_CRANE LIFT"
   Button "Button_2" at 80,238 size 96x32; TextOff 'Left'; Authorization "Maintenance"
      on Press: InvertBit("DB_HMI_CRANE LEFT")
      Appearance <- "DB_HMI_CRANE LEFT"
   Button "Button_3" at 80,279 size 96x32; TextOff 'Right'; Authorization "Maintenance"
      on Press: InvertBit("DB_HMI_CRANE RIGHT")
      Appearance <- "DB_HMI_CRANE RIGHT"
   Button "Button_4" at 344,198 size 106x32; TextOff 'Rotate CW'; Authorization "Maintenance"
      on Press: InvertBit("DB_HMI_ASSEMPLER ROT CW")
      Appearance <- "DB_HMI_ASSEMPLER ROT CW"
   Button "Button_5" at 345,238 size 104x32; TextOff 'Rotate CCW'; Authorization "Maintenance"
      on Press: InvertBit("DB_HMI_ASSEMPLER ROT CCW")
      Appearance <- "DB_HMI_ASSEMPLER ROT CCW"
   Button "Button_6" at 346,279 size 103x32; TextOff 'Grab'; Authorization "Maintenance"
      on Press: InvertBit("DB_HMI_ASSEMPLER GRAB")
      Appearance <- "DB_HMI_ASSEMPLER GRAB"
   TextField "Text field_5" at 303,119 size 82x23; Text 'X Target:'
   TextField "Text field_6" at 302,159 size 81x23; Text 'Z Target:'
   IOField "I/O field_3" at 397,110 size 96x32; Authorization "Maintenance"; FormatPattern 99.999
      ProcessValue <- "DB_HMI_ASSEMPLER X"
   IOField "I/O field_4" at 397,150 size 96x32; Authorization "Maintenance"; FormatPattern 99.999
      ProcessValue <- "DB_HMI_ASSEMPLER Z"
   TextField "Text field_7" at 641,62 size 84x32; Text 'Resets'
   Button "Button_7" at 597,110 size 173x32; TextOff 'Rack Memory Reset'; Authorization "Maintenance"
      on Press: SetBit("DB_RackMemory_ReckMemoryReset")
   Button "Button_8" at 597,150 size 172x32; TextOff 'In Production Reset'; Authorization "Maintenance"
      on Press: SetBit("DB_RackMemory_InProductionReset")
   TextField "Text field_8" at 259,336 size 268x61; Text '*PLEASE MAKE SURE TO RESET THE ASSEMPLER ROTATION TO INITIAL STATE'
   Button "Button_9" at 11,10 size 96x32; TextOff 'LOG IN'
      on Release: function_f41c6f6c("CURRENT USER")
      on Press: function_a2a04561()
   Button "Button_10" at 126,8 size 96x32; TextOff 'LOG OUT'
      on Press: function_f23ef4c9(); SetTag("CURRENT USER", '""')
   Switch "Switch_1" at 159,348 size 64x32; CaptionText 'Switch'; TextOff 'OFF'; TextOn 'ON'; Authorization "Maintenance"
      on SwitchOn: SetBit("DB_HMI_MAINTENANCE MODE")
      on SwitchOff: ResetBit("DB_HMI_MAINTENANCE MODE")
      ProcessValue <- "DB_HMI_MAINTENANCE MODE"
   TextField "Text field_10" at 37,357 size 110x23; Text 'maintenance'
   IOField "I/O field_13" at 685,3 size 106x32; FormatPattern ??????????????????????????????????????????????????????????????????????
      ProcessValue <- "CURRENT USER"
   TextField "Text field_9" at 542,8 size 140x23; Text 'CURRENT USER:'

screen "Overview" 800x480
   TextField "HmiScreenItemData" at 313,1 size 176x47; Text 'Overview'
   Circle "Circle_1" at 376,88 size 48x48
      Appearance <- "DB_HMI_FACTORY STATUS"
   TextField "Text field_1" at 329,61 size 143x27; Text 'Factory Status'
   TextField "Text field_3" at 389,179 size 25x23; Text 'Z1'
   TextField "Text field_4" at 622,175 size 25x23; Text 'Z2'
   TextField "Text field_5" at 358,211 size 87x42; Text 'Z3 BUFFER-A'
   TextField "Text field_6" at 604,267 size 61x42; Text 'Z4 UPPER'
   TextField "Text field_7" at 622,327 size 25x23; Text 'Z5'
   TextField "Text field_8" at 36,180 size 121x23; Text 'In Production:'
   TextField "Text field_9" at 36,219 size 150x23; Text 'Items in Buffer A:'
   TextField "Text field_10" at 36,264 size 149x23; Text 'Items in Buffer B:'
   TextField "Text field_13" at 36,307 size 145x23; Text 'Occupied Spaces:'
   Bar "Bar_1" at 31,339 size 275x33; MinimumValue 0; MaximumValue 108
      ProcessValue <- "DB_RackMemory_SpacesOccupied"
   Button "Button_12" at 69,415 size 163x52; TextOff 'Production'; Authorization "Operate"
      on Release: ActivateScreen("Production", 0)
   Button "Button_13" at 238,415 size 163x52; TextOff 'Warehouse'
      on Release: ActivateScreen("Warehouse", 0)
   Button "Button_14" at 408,415 size 163x52; TextOff 'Alarms'
      on Release: ActivateScreen("Alarms", 0)
   Button "Button_15" at 578,415 size 163x52; TextOff 'Maintenance'; Authorization "Maintenance"
      on Release: ActivateScreen("Maintenance", 0)
   IOField "I/O field_1" at 202,176 size 96x32; FormatPattern 99
      ProcessValue <- "DB_RackMemory_In_Production"
   IOField "I/O field_4" at 203,215 size 96x32; FormatPattern 99
      ProcessValue <- "ZONE-3 BUFFER_A_DB_BUFFER_ITEMS_COUNT_CV"
   IOField "I/O field_5" at 203,260 size 96x32; FormatPattern 99
      ProcessValue <- "Zone_3_FB_DB_ZONE-3 BUFFER B_BUFFER_ITEMS_COUNT_CV"
   IOField "I/O field_6" at 203,303 size 96x32; FormatPattern 999
      ProcessValue <- "DB_RackMemory_SpacesOccupied"
   IOField "I/O field_7" at 452,175 size 96x32; FormatPattern 999
      ProcessValue <- "DB_HMI_Z1 STATUS"
   IOField "I/O field_8" at 680,173 size 96x32; FormatPattern 999
      ProcessValue <- "DB_HMI_Z2 STATUS"
   IOField "I/O field_9" at 680,273 size 96x32; FormatPattern 999
      ProcessValue <- "DB_HMI_Z4 UPPER STATUS"
   IOField "I/O field_10" at 452,226 size 96x32; FormatPattern 999
      ProcessValue <- "DB_HMI_Z3 BUFFER A STATUS"
   IOField "I/O field_11" at 680,324 size 96x32; FormatPattern 999
      ProcessValue <- "DB_HMI_Z5 STATUS"
   TextField "Text field_11" at 592,220 size 86x42; Text 'Z3 BUFFER-B'
   IOField "I/O field_2" at 680,223 size 96x32; FormatPattern 999
      ProcessValue <- "DB_HMI_Z3 BUFFER B STATUS"
   TextField "Text field_12" at 348,264 size 103x42; Text 'Z3 ASSEMPLER'
   IOField "I/O field_3" at 452,274 size 96x32; FormatPattern 999
      ProcessValue <- "DB_HMI_Z3 ASSEMPLER STATUS"
   TextField "Text field_14" at 370,315 size 64x42; Text 'Z4 LOWER'
   IOField "I/O field_12" at 452,326 size 96x32; FormatPattern 999
      ProcessValue <- "DB_HMI_Z4 LOWER STATUS"
   Button "Button_1" at 11,10 size 96x32; TextOff 'LOG IN'
      on Press: function_a2a04561()
      on Release: function_f41c6f6c("CURRENT USER")
   Button "Button_2" at 126,8 size 96x32; TextOff 'LOG OUT'
      on Press: function_f23ef4c9(); SetTag("CURRENT USER", '""')
   IOField "I/O field_13" at 685,3 size 106x32; FormatPattern ??????????????????????????????????????????????????????????????????????
      ProcessValue <- "CURRENT USER"
   TextField "Text field_2" at 542,8 size 140x23; Text 'CURRENT USER:'
*)